VERSION : 0.1
   VAR
      "1#排气阀关到位" : Bool;
      "1#排气阀开到位" : Bool;
      "1#进料阀关到位" : Bool;
      "1#进料阀开到位" : Bool;
      "1#出料阀关到位" : Bool;
      "1#出料阀开到位" : Bool;
      "1#进气阀关到位" : Bool;
      "1#进气阀开到位" : Bool;
      "1#助吹阀关到位" : Bool;
      "1#助吹阀开到位" : Bool;
      "1#排堵阀关到位" : Bool;
      "1#排堵阀开到位" : Bool;
      "1#料位信号" : Bool;
      "1#现场箱远程" : Bool;
      "2#排气阀关到位" : Bool;
      "2#排气阀开到位" : Bool;
      "2#进料阀关到位" : Bool;
      "2#进料阀开到位" : Bool;
      "2#出料阀关到位" : Bool;
      "2#出料阀开到位" : Bool;
      "2#进气阀关到位" : Bool;
      "2#进气阀开到位" : Bool;
      "2#助吹阀关到位" : Bool;
      "2#助吹阀开到位" : Bool;
      "2#排堵阀关到位" : Bool;
      "2#排堵阀开到位" : Bool;
      "2#料位信号" : Bool;
      "2#现场箱远程" : Bool;
      "1#切1#切换阀关到位" : Bool;
      "1#切1#切换阀开到位" : Bool;
      "1#切2#切换阀关到位" : Bool;
      "1#切2#切换阀开到位" : Bool;
      "1#切3#切换阀关到位" : Bool;
      "1#切3#切换阀开到位" : Bool;
      "1#切4#切换阀关到位" : Bool;
      "1#切4#切换阀开到位" : Bool;
      "1#切5#切换阀关到位" : Bool;
      "1#切5#切换阀开到位" : Bool;
      "1#切远程信号" : Bool;
      "2#切1#切换阀关到位" : Bool;
      "2#切1#切换阀开到位" : Bool;
      "2#切2#切换阀关到位" : Bool;
      "2#切2#切换阀开到位" : Bool;
      "2#切远程信号" : Bool;
      "3#切1#切换阀关到位" : Bool;
      "3#切1#切换阀开到位" : Bool;
      "3#切2#切换阀关到位" : Bool;
      "3#切2#切换阀开到位" : Bool;
      "3#切远程信号" : Bool;
      "4#切1#切换阀关到位" : Bool;
      "4#切1#切换阀开到位" : Bool;
      "4#切2#切换阀关到位" : Bool;
      "4#切2#切换阀开到位" : Bool;
      "4#切3#切换阀关到位" : Bool;
      "4#切3#切换阀开到位" : Bool;
      "4#切4#切换阀关到位" : Bool;
      "4#切4#切换阀开到位" : Bool;
      "4#切远程信号" : Bool;
      "1#中控备妥" : Bool;
      "1#运行" : Bool;
      "1#母管压力低" : Bool;
      "1#灰管压力高" : Bool;
      "2#中控备妥" : Bool;
      "2#运行" : Bool;
      "2#母管压力低" : Bool;
      "2#灰管压力高" : Bool;
      STAT66 : Bool;
      STAT67 : Bool;
      STAT68 : Bool;
      STAT69 : Bool;
      STAT70 : Bool;
      STAT71 : Bool;
      STAT72 : Bool;
      STAT73 : Bool;
      STAT74 : Bool;
      STAT75 : Bool;
      STAT76 : Bool;
      STAT77 : Bool;
      STAT78 : Bool;
      STAT79 : Bool;
      STAT80 : Bool;
      STAT81 : Bool;
      STAT82 : Bool;
      STAT83 : Bool;
      STAT84 : Bool;
      STAT85 : Bool;
      STAT86 : Bool;
      STAT87 : Bool;
      STAT88 : Bool;
      STAT89 : Bool;
      STAT90 : Bool;
      STAT91 : Bool;
      STAT92 : Bool;
      STAT93 : Bool;
      STAT94 : Bool;
      STAT95 : Bool;
      STAT96 : Bool;
      STAT97 : Bool;
      STAT98 : Bool;
      STAT99 : Bool;
      STAT100 : Bool;
      STAT101 : Bool;
      STAT102 : Bool;
      STAT103 : Bool;
      STAT104 : Bool;
      STAT105 : Bool;
      STAT106 : Bool;
      STAT107 : Bool;
      STAT108 : Bool;
      STAT109 : Bool;
      STAT110 : Bool;
      STAT111 : Bool;
      STAT112 : Bool;
      STAT113 : Bool;
      STAT114 : Bool;
      STAT115 : Bool;
      STAT116 : Bool;
      STAT117 : Bool;
      STAT118 : Bool;
      STAT119 : Bool;
      STAT120 : Bool;
      STAT121 : Bool;
      STAT122 : Bool;
      STAT123 : Bool;
      STAT124 : Bool;
      STAT125 : Bool;
      STAT126 : Bool;
      STAT127 : Bool;
      STAT128 : Bool;
      STAT129 : Bool;
      STAT130 : Bool;
      STAT131 : Bool;
      STAT132 : Bool;
      STAT133 : Bool;
      STAT134 : Bool;
      STAT135 : Bool;
      STAT136 : Bool;
      STAT137 : Bool;
      STAT138 : Bool;
      STAT139 : Bool;
      STAT140 : Bool;
      STAT141 : Bool;
      STAT142 : Bool;
      STAT143 : Bool;
      STAT144 : Bool;
   END_VAR
BEGIN
END_DATA_BLOCK

DATA_BLOCK "DB20"   // DB20
{ S7_Optimized_Access := 'FALSE' }
VERSION : 0.1
   VAR
      STAT0 : Real;
      STAT1 : Real;
      STAT2 : Real;
      STAT3 : Real;
      STAT4 : Real;
      STAT5 : Real;
      STAT6 : Real;
      STAT7 : Real;
      STAT8 : Real;
      STAT9 : Real;
      STAT10 : Real;
      STAT11 : Real;
      STAT12 : Real;
      STAT13 : Real;
      STAT14 : Real;
      STAT15 : Real;
      STAT16 : Real;
      STAT17 : Real;
      STAT18 : Real;
      STAT19 : Real;
      STAT20 : Real;
      STAT21 : Real;
      STAT22 : Real;
      STAT23 : Real;
      STAT24 : Bool;
      STAT25 : Bool;
      STAT26 : Word;
   END_VAR
BEGIN
END_DATA_BLOCK

FUNCTION_BLOCK "累计功能块"   // FB1, LAD
{ S7_Optimized_Access := 'FALSE' }
VERSION : 0.1
   VAR_INPUT
      CLEAR : Bool;   // 清零
      DATA : Real;   // 瞬时量
   END_VAR
   VAR_OUTPUT
      OUT1 : Real;
   END_VAR
   VAR
      STAT2 : Real;
      STAT3 : Real;
      STAT4 : Real;
      P1 : Bool;
   END_VAR
   VAR_TEMP   // added for the SCL form of the ladder/FBD networks
      _w1 : Bool;
   END_VAR
BEGIN

REGION Network 1
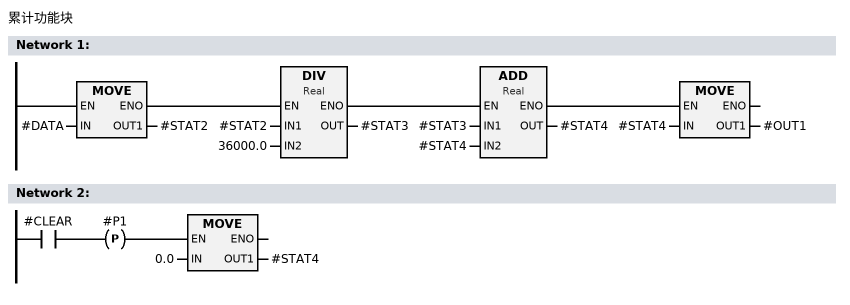
   RUNG wire#powerrail
      { S7_GenerateENO := "TRUE" } Move(in := #DATA, out1 => #STAT2)
      { S7_Templates := "SrcType := Real"; S7_GenerateENO := "TRUE" } Div(in1 := #STAT2, in2 := 36000.0, out => #STAT3)
      { S7_Templates := "SrcType := Real"; S7_GenerateENO := "TRUE" } Add(in1 := #STAT3, in2 := #STAT4, out => #STAT4)
      { S7_GenerateENO := "TRUE" } Move(in := #STAT4, out1 => #OUT1)
   END_RUNG
   // the same network as SCL:
   // ENO of a box is taken as its EN; it also drops when the box reports an error
   #STAT2 := #DATA;
   #STAT3 := #STAT2 / 36000.0;
   #STAT4 := #STAT3 + #STAT4;
   #OUT1 := #STAT4;
END_REGION

REGION Network 2
   RUNG wire#powerrail
      Contact( #CLEAR )
      P_Trig( #P1 )
      { S7_GenerateENO := "TRUE" } Move(in := 0.0, out1 => #STAT4)
   END_RUNG
   // the same network as SCL:
   #_w1 := #CLEAR AND NOT #P1;   // rising edge
   #P1 := #CLEAR;
   IF #_w1 THEN #STAT4 := 0.0; END_IF;
END_REGION
END_FUNCTION_BLOCK

FUNCTION_BLOCK "FB11_DATA_ALARM_FB"   // FB11, LAD
{ S7_Optimized_Access := 'FALSE' }
VERSION : 0.1
   VAR
      PIW256 : "FB330_DATA_ALARM";
      PIW258 : "FB330_DATA_ALARM";
      PIW260 : "FB330_DATA_ALARM";
      PIW262 : "FB330_DATA_ALARM";
      PIW264 : "FB330_DATA_ALARM";
      PIW266 : "FB330_DATA_ALARM";
      PIW268 : "FB330_DATA_ALARM";
      PIW270 : "FB330_DATA_ALARM";
      PIW272 : "FB330_DATA_ALARM";
      PIW274 : "FB330_DATA_ALARM";
      PIW276 : "FB330_DATA_ALARM";
      PIW278 : "FB330_DATA_ALARM";
      PIW280 : "FB330_DATA_ALARM";
      PIW282 : "FB330_DATA_ALARM";
      PIW284 : "FB330_DATA_ALARM";
      PIW286 : "FB330_DATA_ALARM";
      PIW288 : "FB330_DATA_ALARM";
      PIW290 : "FB330_DATA_ALARM";
      PIW292 : "FB330_DATA_ALARM";
      PIW294 : "FB330_DATA_ALARM";
      PIW296 : "FB330_DATA_ALARM";
      PIW298 : "FB330_DATA_ALARM";
      PIW300 : "FB330_DATA_ALARM";
      PIW302 : "FB330_DATA_ALARM";
      PID304 : "FB330_DATA_ALARM";
      PID308 : "FB330_DATA_ALARM";
      PID312 : "FB330_DATA_ALARM";
      PID316 : "FB330_DATA_ALARM";
      PID320 : "FB330_DATA_ALARM";
      PID324 : "FB330_DATA_ALARM";
      PID328 : "FB330_DATA_ALARM";
      PID332 : "FB330_DATA_ALARM";
      PID336 : "FB330_DATA_ALARM";
      PID340 : "FB330_DATA_ALARM";
      PID344 : "FB330_DATA_ALARM";
      PID348 : "FB330_DATA_ALARM";
      PID352 : "FB330_DATA_ALARM";
      PID356 : "FB330_DATA_ALARM";
      PID360 : "FB330_DATA_ALARM";
      PID364 : "FB330_DATA_ALARM";
      PID368 : "FB330_DATA_ALARM";
      PID372 : "FB330_DATA_ALARM";
      PID376 : "FB330_DATA_ALARM";
      PID380 : "FB330_DATA_ALARM";
      PID384 : "FB330_DATA_ALARM";
      PID388 : "FB330_DATA_ALARM";
      PID392 : "FB330_DATA_ALARM";
      PID396 : "FB330_DATA_ALARM";
      IW110 : "FB330_DATA_ALARM";
      IW112 : "FB330_DATA_ALARM";
      IW114 : "FB330_DATA_ALARM";
      IW116 : "FB330_DATA_ALARM";
      PID400 : "FB330_DATA_ALARM";
      PID408 : "FB330_DATA_ALARM";
      PID416 : "FB330_DATA_ALARM";
      Static4 : "FB330_DATA_ALARM";
      Static5 : "FB330_DATA_ALARM";
      Static6 : "FB330_DATA_ALARM";
      Static7 : "FB330_DATA_ALARM";
      Static8 : "FB330_DATA_ALARM";
      Static9 : "FB330_DATA_ALARM";
      Static10 : "FB330_DATA_ALARM";
   END_VAR
BEGIN

REGION Network 1
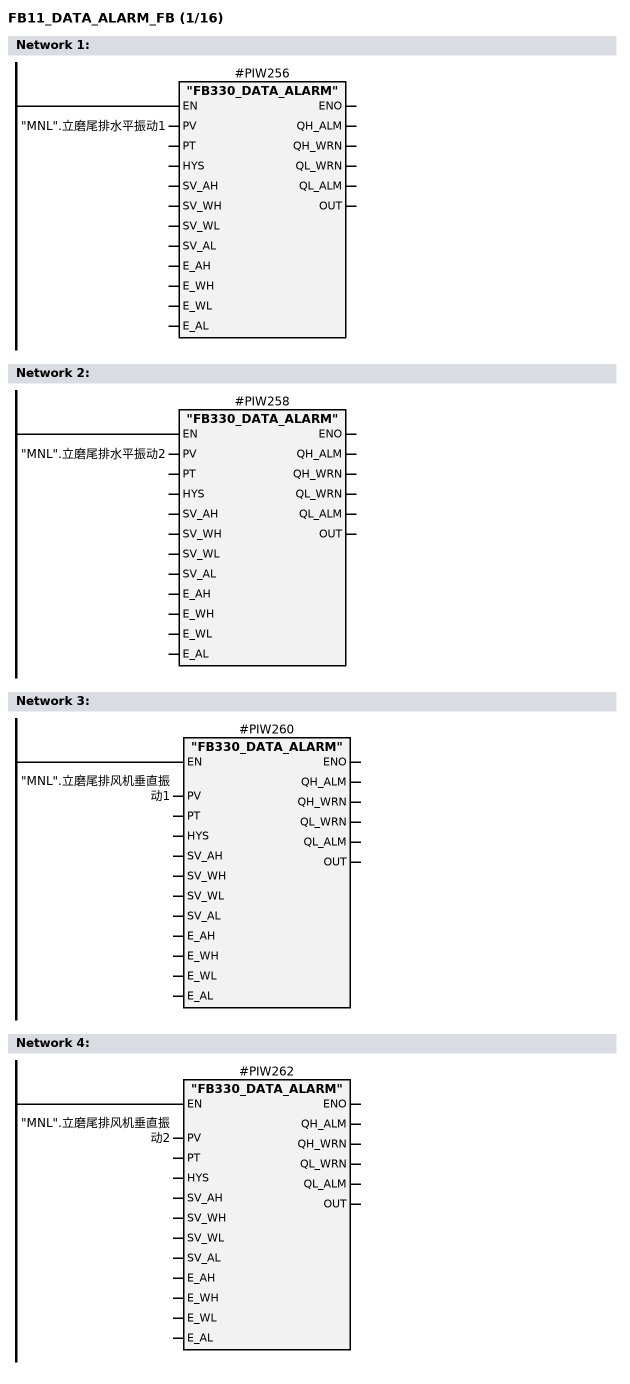
   RUNG wire#powerrail
      #PIW256(PV := "MNL".立磨尾排水平振动1, PT :=, HYS :=, SV_AH :=, SV_WH :=, SV_WL :=, SV_AL :=, E_AH :=, E_WH :=, E_WL :=, E_AL :=, QH_ALM =>, QH_WRN =>, QL_WRN =>, QL_ALM =>, OUT =>)
   END_RUNG
   // the same network as SCL:
   #PIW256(PV := "MNL".立磨尾排水平振动1);   // "FB330_DATA_ALARM"
END_REGION

REGION Network 2
   RUNG wire#powerrail
      #PIW258(PV := "MNL".立磨尾排水平振动2, PT :=, HYS :=, SV_AH :=, SV_WH :=, SV_WL :=, SV_AL :=, E_AH :=, E_WH :=, E_WL :=, E_AL :=, QH_ALM =>, QH_WRN =>, QL_WRN =>, QL_ALM =>, OUT =>)
   END_RUNG
   // the same network as SCL:
   #PIW258(PV := "MNL".立磨尾排水平振动2);   // "FB330_DATA_ALARM"
END_REGION

REGION Network 3
   RUNG wire#powerrail
      #PIW260(PV := "MNL".立磨尾排风机垂直振动1, PT :=, HYS :=, SV_AH :=, SV_WH :=, SV_WL :=, SV_AL :=, E_AH :=, E_WH :=, E_WL :=, E_AL :=, QH_ALM =>, QH_WRN =>, QL_WRN =>, QL_ALM =>, OUT =>)
   END_RUNG
   // the same network as SCL:
   #PIW260(PV := "MNL".立磨尾排风机垂直振动1);   // "FB330_DATA_ALARM"
END_REGION

REGION Network 4
   RUNG wire#powerrail
      #PIW262(PV := "MNL".立磨尾排风机垂直振动2, PT :=, HYS :=, SV_AH :=, SV_WH :=, SV_WL :=, SV_AL :=, E_AH :=, E_WH :=, E_WL :=, E_AL :=, QH_ALM =>, QH_WRN =>, QL_WRN =>, QL_ALM =>, OUT =>)
   END_RUNG
   // the same network as SCL:
   #PIW262(PV := "MNL".立磨尾排风机垂直振动2);   // "FB330_DATA_ALARM"
END_REGION

REGION Network 5
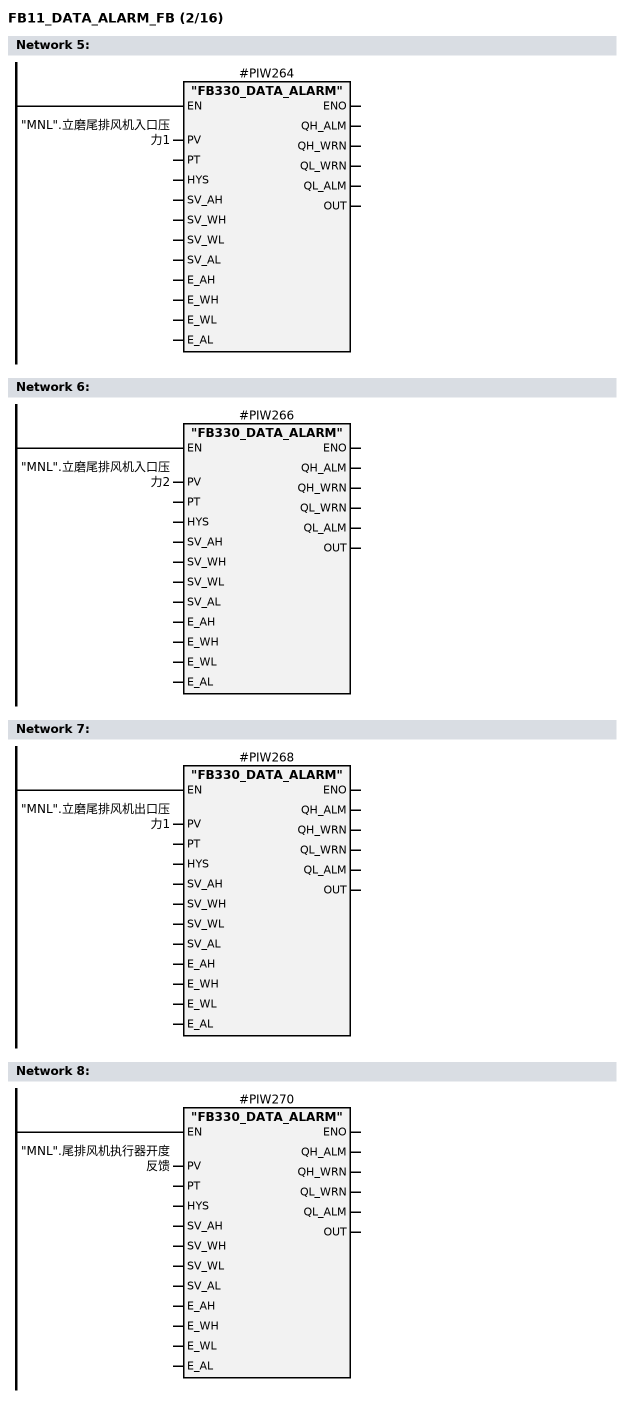
   RUNG wire#powerrail
      #PIW264(PV := "MNL".立磨尾排风机入口压力1, PT :=, HYS :=, SV_AH :=, SV_WH :=, SV_WL :=, SV_AL :=, E_AH :=, E_WH :=, E_WL :=, E_AL :=, QH_ALM =>, QH_WRN =>, QL_WRN =>, QL_ALM =>, OUT =>)
   END_RUNG
   // the same network as SCL:
   #PIW264(PV := "MNL".立磨尾排风机入口压力1);   // "FB330_DATA_ALARM"
END_REGION

REGION Network 6
   RUNG wire#powerrail
      #PIW266(PV := "MNL".立磨尾排风机入口压力2, PT :=, HYS :=, SV_AH :=, SV_WH :=, SV_WL :=, SV_AL :=, E_AH :=, E_WH :=, E_WL :=, E_AL :=, QH_ALM =>, QH_WRN =>, QL_WRN =>, QL_ALM =>, OUT =>)
   END_RUNG
   // the same network as SCL:
   #PIW266(PV := "MNL".立磨尾排风机入口压力2);   // "FB330_DATA_ALARM"
END_REGION

REGION Network 7
   RUNG wire#powerrail
      #PIW268(PV := "MNL".立磨尾排风机出口压力1, PT :=, HYS :=, SV_AH :=, SV_WH :=, SV_WL :=, SV_AL :=, E_AH :=, E_WH :=, E_WL :=, E_AL :=, QH_ALM =>, QH_WRN =>, QL_WRN =>, QL_ALM =>, OUT =>)
   END_RUNG
   // the same network as SCL:
   #PIW268(PV := "MNL".立磨尾排风机出口压力1);   // "FB330_DATA_ALARM"
END_REGION

REGION Network 8
   RUNG wire#powerrail
      #PIW270(PV := "MNL".尾排风机执行器开度反馈, PT :=, HYS :=, SV_AH :=, SV_WH :=, SV_WL :=, SV_AL :=, E_AH :=, E_WH :=, E_WL :=, E_AL :=, QH_ALM =>, QH_WRN =>, QL_WRN =>, QL_ALM =>, OUT =>)
   END_RUNG
   // the same network as SCL:
   #PIW270(PV := "MNL".尾排风机执行器开度反馈);   // "FB330_DATA_ALARM"
END_REGION

REGION Network 9
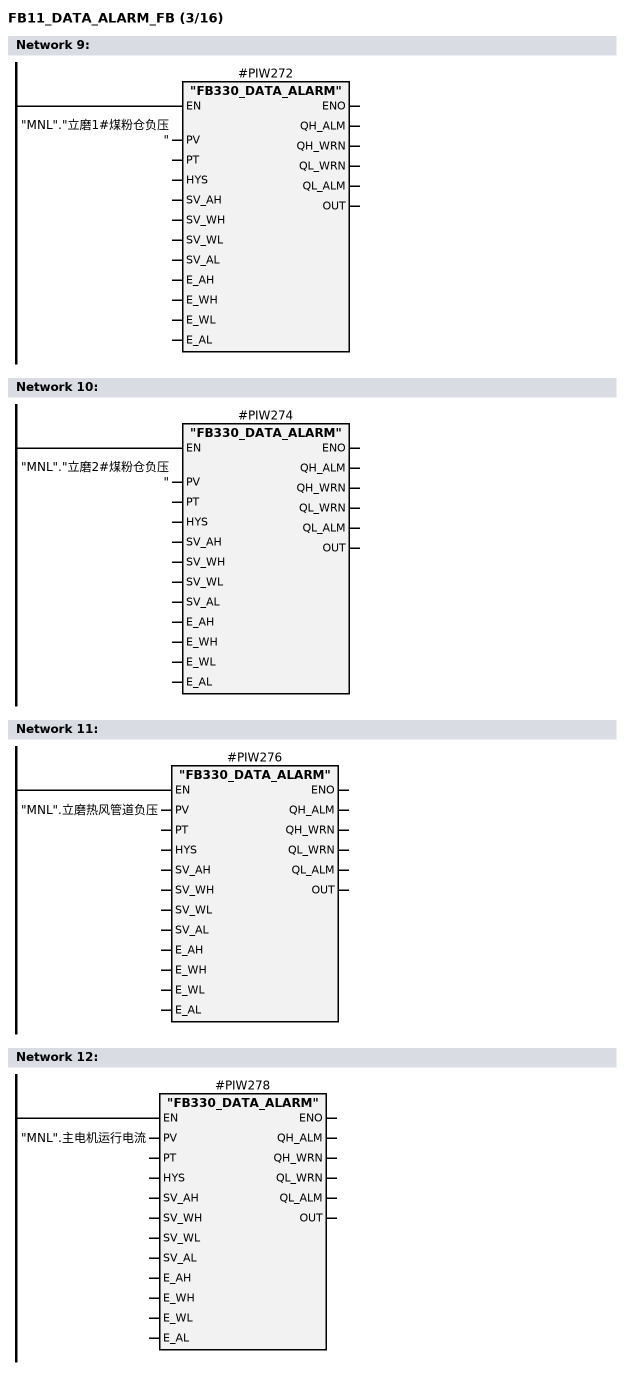
   RUNG wire#powerrail
      #PIW272(PV := "MNL"."立磨1#煤粉仓负压", PT :=, HYS :=, SV_AH :=, SV_WH :=, SV_WL :=, SV_AL :=, E_AH :=, E_WH :=, E_WL :=, E_AL :=, QH_ALM =>, QH_WRN =>, QL_WRN =>, QL_ALM =>, OUT =>)
   END_RUNG
   // the same network as SCL:
   #PIW272(PV := "MNL"."立磨1#煤粉仓负压");   // "FB330_DATA_ALARM"
END_REGION

REGION Network 10
   RUNG wire#powerrail
      #PIW274(PV := "MNL"."立磨2#煤粉仓负压", PT :=, HYS :=, SV_AH :=, SV_WH :=, SV_WL :=, SV_AL :=, E_AH :=, E_WH :=, E_WL :=, E_AL :=, QH_ALM =>, QH_WRN =>, QL_WRN =>, QL_ALM =>, OUT =>)
   END_RUNG
   // the same network as SCL:
   #PIW274(PV := "MNL"."立磨2#煤粉仓负压");   // "FB330_DATA_ALARM"
END_REGION

REGION Network 11
   RUNG wire#powerrail
      #PIW276(PV := "MNL".立磨热风管道负压, PT :=, HYS :=, SV_AH :=, SV_WH :=, SV_WL :=, SV_AL :=, E_AH :=, E_WH :=, E_WL :=, E_AL :=, QH_ALM =>, QH_WRN =>, QL_WRN =>, QL_ALM =>, OUT =>)
   END_RUNG
   // the same network as SCL:
   #PIW276(PV := "MNL".立磨热风管道负压);   // "FB330_DATA_ALARM"
END_REGION

REGION Network 12
   RUNG wire#powerrail
      #PIW278(PV := "MNL".主电机运行电流, PT :=, HYS :=, SV_AH :=, SV_WH :=, SV_WL :=, SV_AL :=, E_AH :=, E_WH :=, E_WL :=, E_AL :=, QH_ALM =>, QH_WRN =>, QL_WRN =>, QL_ALM =>, OUT =>)
   END_RUNG
   // the same network as SCL:
   #PIW278(PV := "MNL".主电机运行电流);   // "FB330_DATA_ALARM"
END_REGION

REGION Network 13
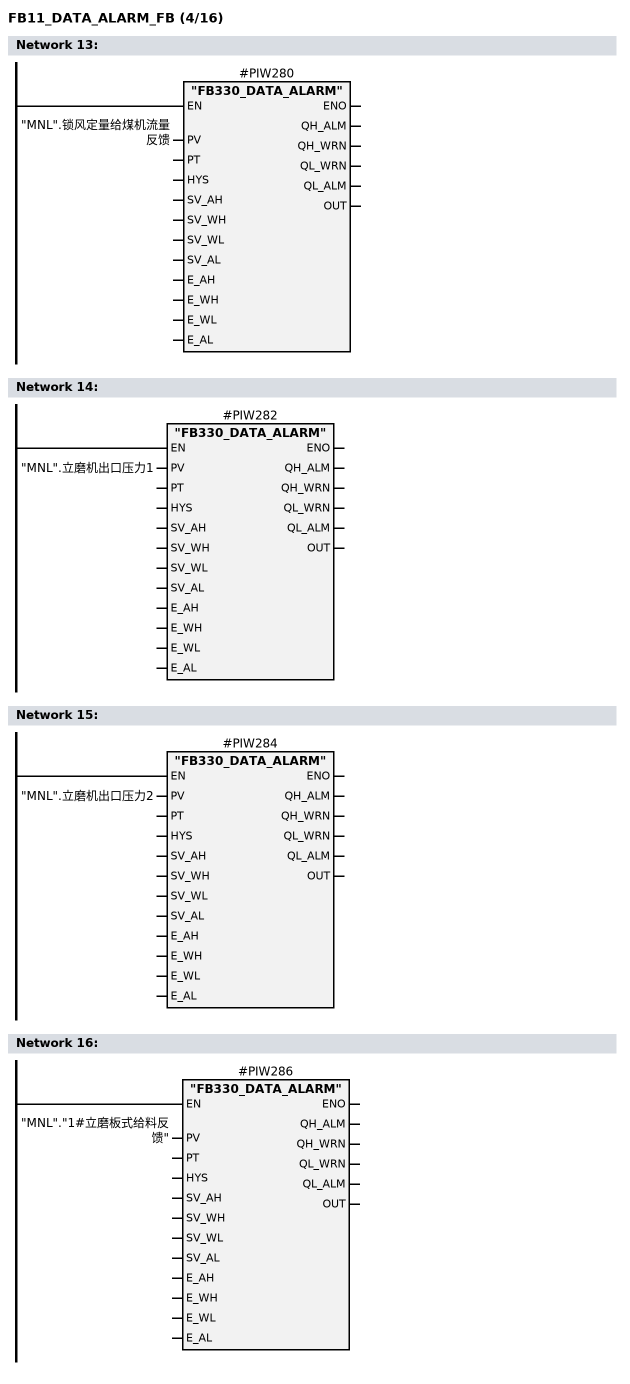
   RUNG wire#powerrail
      #PIW280(PV := "MNL".锁风定量给煤机流量反馈, PT :=, HYS :=, SV_AH :=, SV_WH :=, SV_WL :=, SV_AL :=, E_AH :=, E_WH :=, E_WL :=, E_AL :=, QH_ALM =>, QH_WRN =>, QL_WRN =>, QL_ALM =>, OUT =>)
   END_RUNG
   // the same network as SCL:
   #PIW280(PV := "MNL".锁风定量给煤机流量反馈);   // "FB330_DATA_ALARM"
END_REGION

REGION Network 14
   RUNG wire#powerrail
      #PIW282(PV := "MNL".立磨机出口压力1, PT :=, HYS :=, SV_AH :=, SV_WH :=, SV_WL :=, SV_AL :=, E_AH :=, E_WH :=, E_WL :=, E_AL :=, QH_ALM =>, QH_WRN =>, QL_WRN =>, QL_ALM =>, OUT =>)
   END_RUNG
   // the same network as SCL:
   #PIW282(PV := "MNL".立磨机出口压力1);   // "FB330_DATA_ALARM"
END_REGION

REGION Network 15
   RUNG wire#powerrail
      #PIW284(PV := "MNL".立磨机出口压力2, PT :=, HYS :=, SV_AH :=, SV_WH :=, SV_WL :=, SV_AL :=, E_AH :=, E_WH :=, E_WL :=, E_AL :=, QH_ALM =>, QH_WRN =>, QL_WRN =>, QL_ALM =>, OUT =>)
   END_RUNG
   // the same network as SCL:
   #PIW284(PV := "MNL".立磨机出口压力2);   // "FB330_DATA_ALARM"
END_REGION

REGION Network 16
   RUNG wire#powerrail
      #PIW286(PV := "MNL"."1#立磨板式给料反馈", PT :=, HYS :=, SV_AH :=, SV_WH :=, SV_WL :=, SV_AL :=, E_AH :=, E_WH :=, E_WL :=, E_AL :=, QH_ALM =>, QH_WRN =>, QL_WRN =>, QL_ALM =>, OUT =>)
   END_RUNG
   // the same network as SCL:
   #PIW286(PV := "MNL"."1#立磨板式给料反馈");   // "FB330_DATA_ALARM"
END_REGION

REGION Network 17
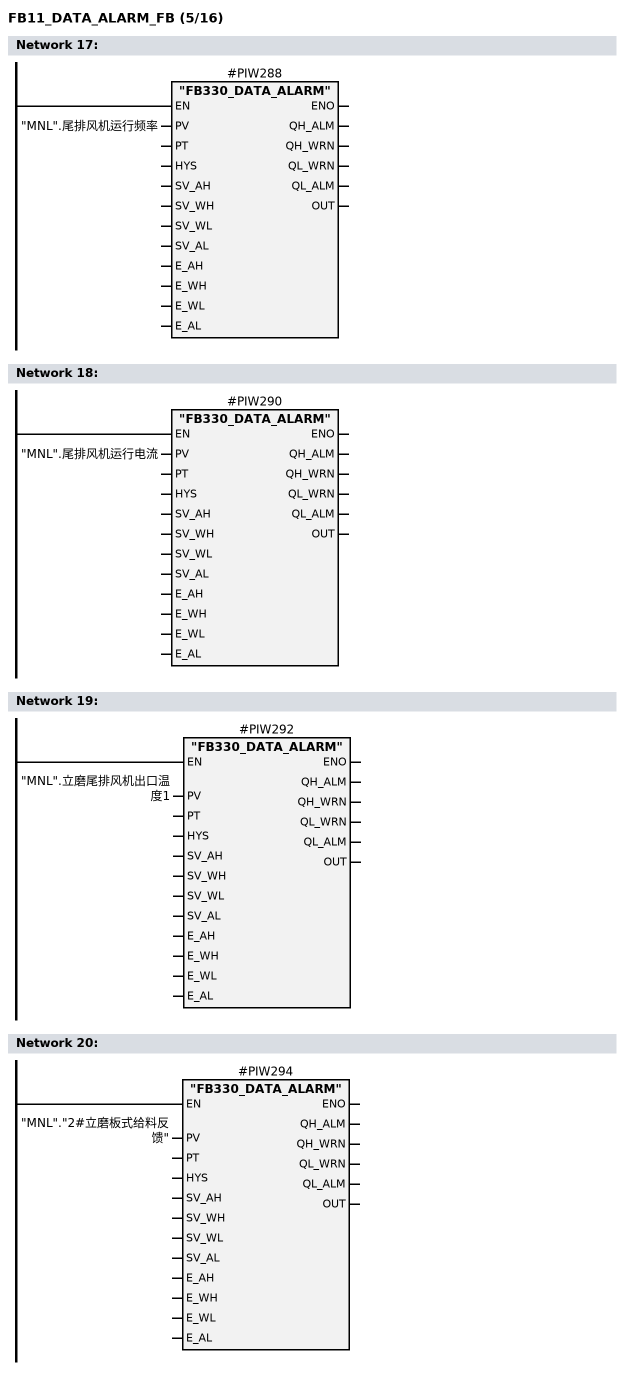
   RUNG wire#powerrail
      #PIW288(PV := "MNL".尾排风机运行频率, PT :=, HYS :=, SV_AH :=, SV_WH :=, SV_WL :=, SV_AL :=, E_AH :=, E_WH :=, E_WL :=, E_AL :=, QH_ALM =>, QH_WRN =>, QL_WRN =>, QL_ALM =>, OUT =>)
   END_RUNG
   // the same network as SCL:
   #PIW288(PV := "MNL".尾排风机运行频率);   // "FB330_DATA_ALARM"
END_REGION

REGION Network 18
   RUNG wire#powerrail
      #PIW290(PV := "MNL".尾排风机运行电流, PT :=, HYS :=, SV_AH :=, SV_WH :=, SV_WL :=, SV_AL :=, E_AH :=, E_WH :=, E_WL :=, E_AL :=, QH_ALM =>, QH_WRN =>, QL_WRN =>, QL_ALM =>, OUT =>)
   END_RUNG
   // the same network as SCL:
   #PIW290(PV := "MNL".尾排风机运行电流);   // "FB330_DATA_ALARM"
END_REGION

REGION Network 19
   RUNG wire#powerrail
      #PIW292(PV := "MNL".立磨尾排风机出口温度1, PT :=, HYS :=, SV_AH :=, SV_WH :=, SV_WL :=, SV_AL :=, E_AH :=, E_WH :=, E_WL :=, E_AL :=, QH_ALM =>, QH_WRN =>, QL_WRN =>, QL_ALM =>, OUT =>)
   END_RUNG
   // the same network as SCL:
   #PIW292(PV := "MNL".立磨尾排风机出口温度1);   // "FB330_DATA_ALARM"
END_REGION

REGION Network 20
   RUNG wire#powerrail
      #PIW294(PV := "MNL"."2#立磨板式给料反馈", PT :=, HYS :=, SV_AH :=, SV_WH :=, SV_WL :=, SV_AL :=, E_AH :=, E_WH :=, E_WL :=, E_AL :=, QH_ALM =>, QH_WRN =>, QL_WRN =>, QL_ALM =>, OUT =>)
   END_RUNG
   // the same network as SCL:
   #PIW294(PV := "MNL"."2#立磨板式给料反馈");   // "FB330_DATA_ALARM"
END_REGION

REGION Network 21
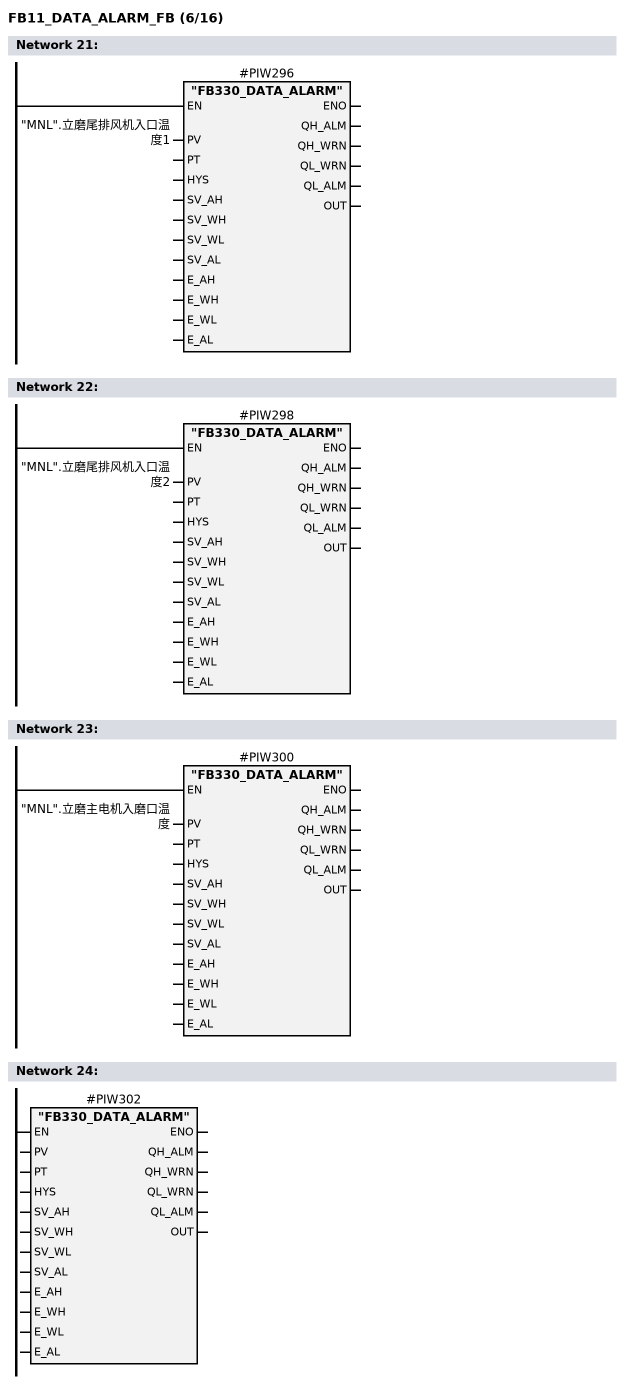
   RUNG wire#powerrail
      #PIW296(PV := "MNL".立磨尾排风机入口温度1, PT :=, HYS :=, SV_AH :=, SV_WH :=, SV_WL :=, SV_AL :=, E_AH :=, E_WH :=, E_WL :=, E_AL :=, QH_ALM =>, QH_WRN =>, QL_WRN =>, QL_ALM =>, OUT =>)
   END_RUNG
   // the same network as SCL:
   #PIW296(PV := "MNL".立磨尾排风机入口温度1);   // "FB330_DATA_ALARM"
END_REGION

REGION Network 22
   RUNG wire#powerrail
      #PIW298(PV := "MNL".立磨尾排风机入口温度2, PT :=, HYS :=, SV_AH :=, SV_WH :=, SV_WL :=, SV_AL :=, E_AH :=, E_WH :=, E_WL :=, E_AL :=, QH_ALM =>, QH_WRN =>, QL_WRN =>, QL_ALM =>, OUT =>)
   END_RUNG
   // the same network as SCL:
   #PIW298(PV := "MNL".立磨尾排风机入口温度2);   // "FB330_DATA_ALARM"
END_REGION

REGION Network 23
   RUNG wire#powerrail
      #PIW300(PV := "MNL".立磨主电机入磨口温度, PT :=, HYS :=, SV_AH :=, SV_WH :=, SV_WL :=, SV_AL :=, E_AH :=, E_WH :=, E_WL :=, E_AL :=, QH_ALM =>, QH_WRN =>, QL_WRN =>, QL_ALM =>, OUT =>)
   END_RUNG
   // the same network as SCL:
   #PIW300(PV := "MNL".立磨主电机入磨口温度);   // "FB330_DATA_ALARM"
END_REGION

REGION Network 24
   RUNG wire#powerrail
      #PIW302(PV :=, PT :=, HYS :=, SV_AH :=, SV_WH :=, SV_WL :=, SV_AL :=, E_AH :=, E_WH :=, E_WL :=, E_AL :=, QH_ALM =>, QH_WRN =>, QL_WRN =>, QL_ALM =>, OUT =>)
   END_RUNG
   // the same network as SCL:
   #PIW302();   // "FB330_DATA_ALARM"
END_REGION

REGION Network 25
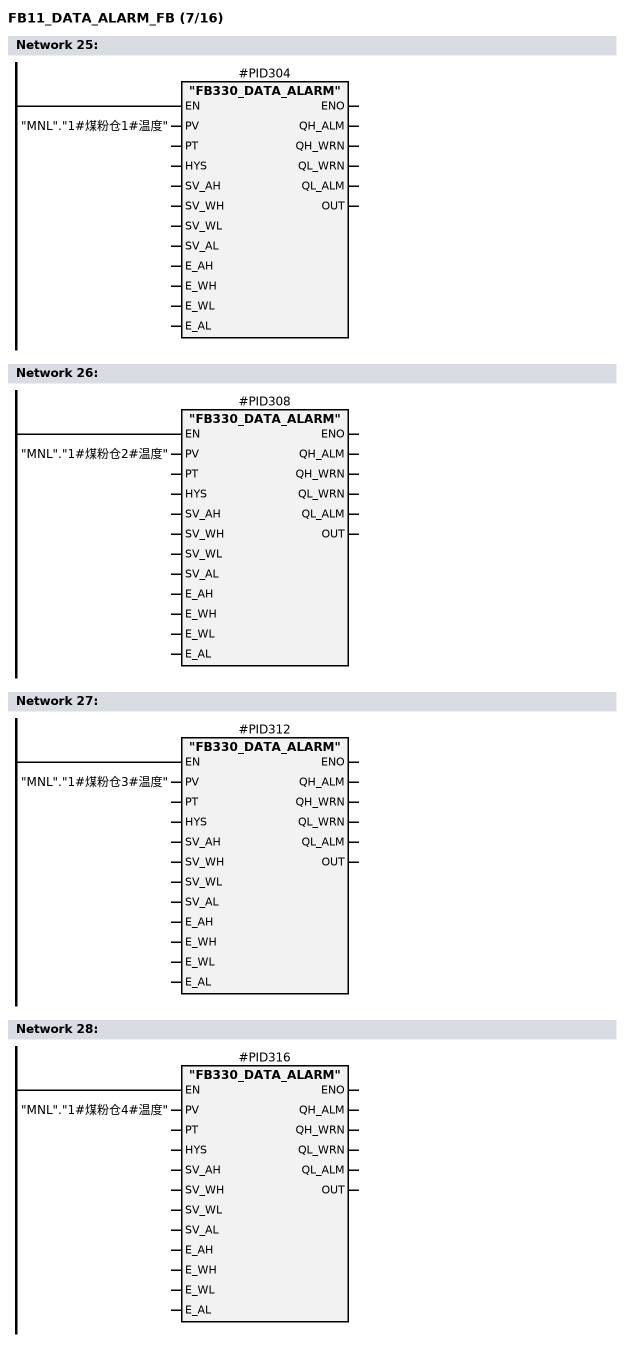
   RUNG wire#powerrail
      #PID304(PV := "MNL"."1#煤粉仓1#温度", PT :=, HYS :=, SV_AH :=, SV_WH :=, SV_WL :=, SV_AL :=, E_AH :=, E_WH :=, E_WL :=, E_AL :=, QH_ALM =>, QH_WRN =>, QL_WRN =>, QL_ALM =>, OUT =>)
   END_RUNG
   // the same network as SCL:
   #PID304(PV := "MNL"."1#煤粉仓1#温度");   // "FB330_DATA_ALARM"
END_REGION

REGION Network 26
   RUNG wire#powerrail
      #PID308(PV := "MNL"."1#煤粉仓2#温度", PT :=, HYS :=, SV_AH :=, SV_WH :=, SV_WL :=, SV_AL :=, E_AH :=, E_WH :=, E_WL :=, E_AL :=, QH_ALM =>, QH_WRN =>, QL_WRN =>, QL_ALM =>, OUT =>)
   END_RUNG
   // the same network as SCL:
   #PID308(PV := "MNL"."1#煤粉仓2#温度");   // "FB330_DATA_ALARM"
END_REGION

REGION Network 27
   RUNG wire#powerrail
      #PID312(PV := "MNL"."1#煤粉仓3#温度", PT :=, HYS :=, SV_AH :=, SV_WH :=, SV_WL :=, SV_AL :=, E_AH :=, E_WH :=, E_WL :=, E_AL :=, QH_ALM =>, QH_WRN =>, QL_WRN =>, QL_ALM =>, OUT =>)
   END_RUNG
   // the same network as SCL:
   #PID312(PV := "MNL"."1#煤粉仓3#温度");   // "FB330_DATA_ALARM"
END_REGION

REGION Network 28
   RUNG wire#powerrail
      #PID316(PV := "MNL"."1#煤粉仓4#温度", PT :=, HYS :=, SV_AH :=, SV_WH :=, SV_WL :=, SV_AL :=, E_AH :=, E_WH :=, E_WL :=, E_AL :=, QH_ALM =>, QH_WRN =>, QL_WRN =>, QL_ALM =>, OUT =>)
   END_RUNG
   // the same network as SCL:
   #PID316(PV := "MNL"."1#煤粉仓4#温度");   // "FB330_DATA_ALARM"
END_REGION

REGION Network 29
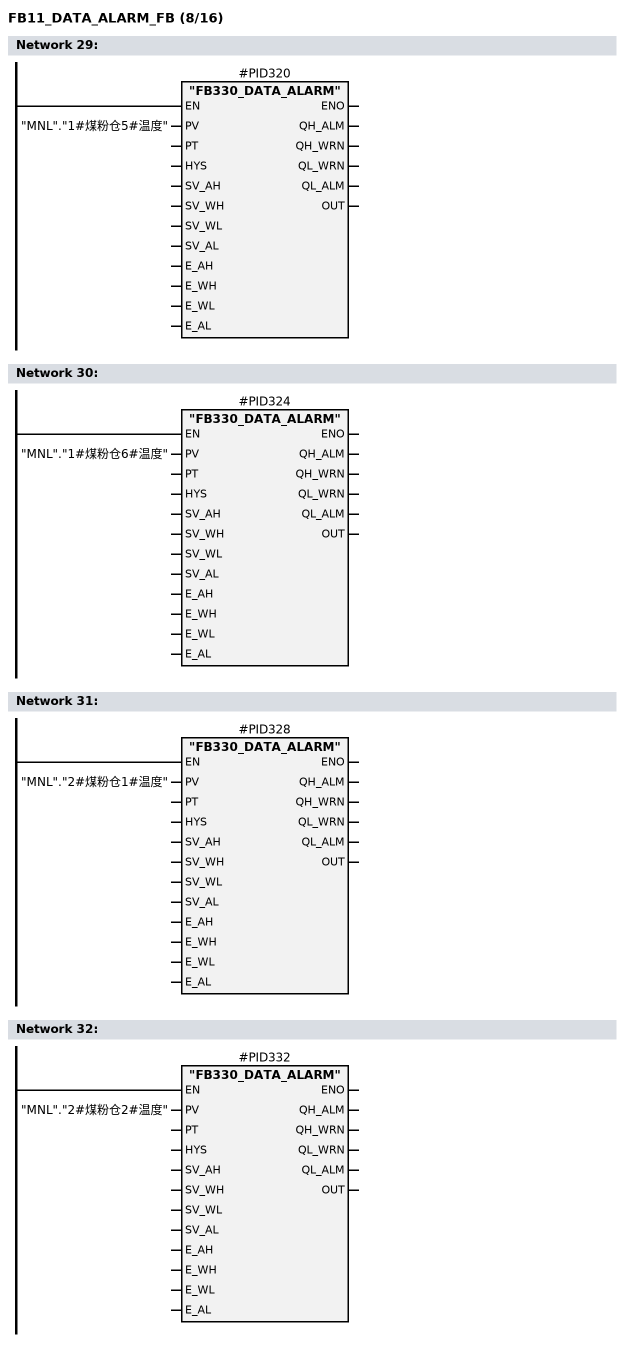
   RUNG wire#powerrail
      #PID320(PV := "MNL"."1#煤粉仓5#温度", PT :=, HYS :=, SV_AH :=, SV_WH :=, SV_WL :=, SV_AL :=, E_AH :=, E_WH :=, E_WL :=, E_AL :=, QH_ALM =>, QH_WRN =>, QL_WRN =>, QL_ALM =>, OUT =>)
   END_RUNG
   // the same network as SCL:
   #PID320(PV := "MNL"."1#煤粉仓5#温度");   // "FB330_DATA_ALARM"
END_REGION

REGION Network 30
   RUNG wire#powerrail
      #PID324(PV := "MNL"."1#煤粉仓6#温度", PT :=, HYS :=, SV_AH :=, SV_WH :=, SV_WL :=, SV_AL :=, E_AH :=, E_WH :=, E_WL :=, E_AL :=, QH_ALM =>, QH_WRN =>, QL_WRN =>, QL_ALM =>, OUT =>)
   END_RUNG
   // the same network as SCL:
   #PID324(PV := "MNL"."1#煤粉仓6#温度");   // "FB330_DATA_ALARM"
END_REGION

REGION Network 31
   RUNG wire#powerrail
      #PID328(PV := "MNL"."2#煤粉仓1#温度", PT :=, HYS :=, SV_AH :=, SV_WH :=, SV_WL :=, SV_AL :=, E_AH :=, E_WH :=, E_WL :=, E_AL :=, QH_ALM =>, QH_WRN =>, QL_WRN =>, QL_ALM =>, OUT =>)
   END_RUNG
   // the same network as SCL:
   #PID328(PV := "MNL"."2#煤粉仓1#温度");   // "FB330_DATA_ALARM"
END_REGION

REGION Network 32
   RUNG wire#powerrail
      #PID332(PV := "MNL"."2#煤粉仓2#温度", PT :=, HYS :=, SV_AH :=, SV_WH :=, SV_WL :=, SV_AL :=, E_AH :=, E_WH :=, E_WL :=, E_AL :=, QH_ALM =>, QH_WRN =>, QL_WRN =>, QL_ALM =>, OUT =>)
   END_RUNG
   // the same network as SCL:
   #PID332(PV := "MNL"."2#煤粉仓2#温度");   // "FB330_DATA_ALARM"
END_REGION

REGION Network 33